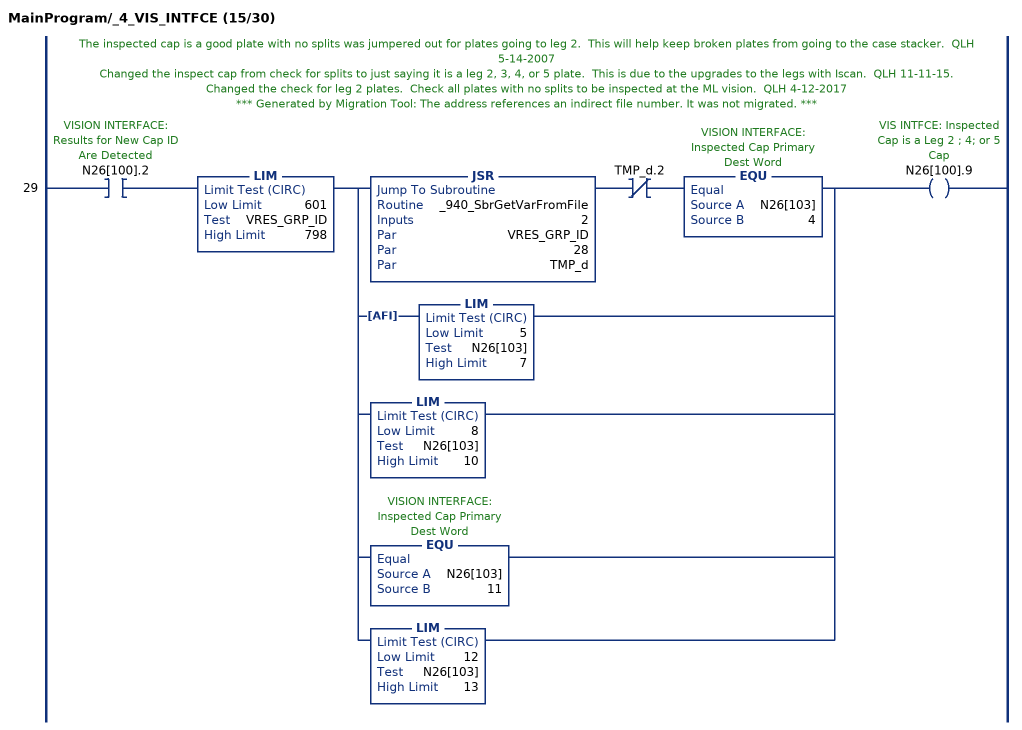
   // The inspected cap is a good plate with no splits was jumpered out for plates going to leg 2.  This will help keep broken plates from going to the case stacker.  QLH 5-14-2007
   // Changed the inspect cap from check for splits to just saying it is a leg 2, 3, 4, or 5 plate.  This is due to the upgrades to the legs with Iscan.  QLH 11-11-15.  Changed the check for leg 2 plates.  Check all plates with no splits to be inspected at the ML vision.  QLH 4-12-2017
   // *** Generated by Migration Tool: The address references an indirect file number. It was not migrated. ***
   29: XIC(N26[100].2)LIM(601,VRES_GRP_ID,798)[JSR(_940_SbrGetVarFromFile,2,VRES_GRP_ID,28,TMP_d) XIO(TMP_d.2) EQU(N26[103],4) ,AFI() LIM(5,N26[103],7) ,LIM(8,N26[103],10) ,EQU(N26[103],11) ,LIM(12,N26[103],13) ]OTE(N26[100].9);
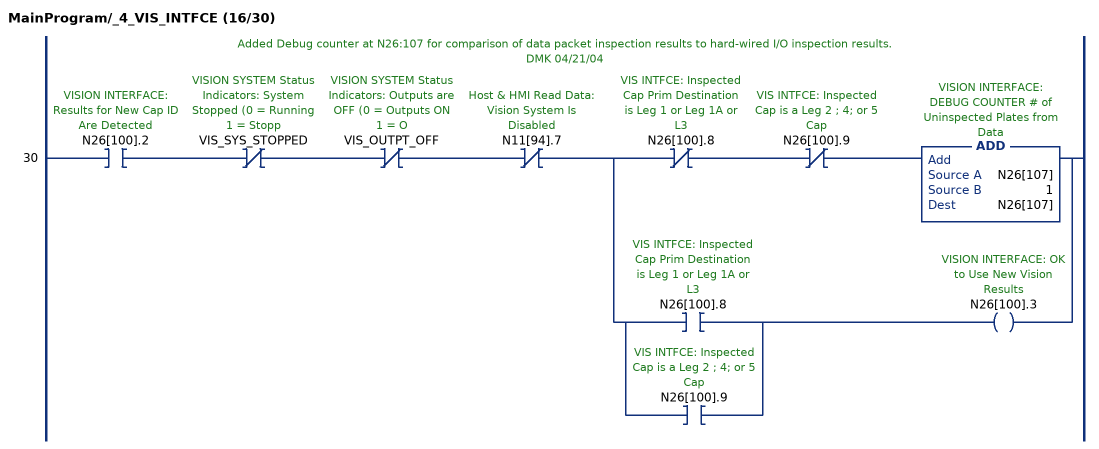
   // Added Debug counter at N26:107 for comparison of data packet inspection results to hard-wired I/O inspection results.
   // DMK 04/21/04
   30: XIC(N26[100].2)XIO(VIS_SYS_STOPPED)XIO(VIS_OUTPT_OFF)XIO(N11[94].7)[XIO(N26[100].8) XIO(N26[100].9) ADD(N26[107],1,N26[107]) ,[XIC(N26[100].8) ,XIC(N26[100].9) ] OTE(N26[100].3) ];
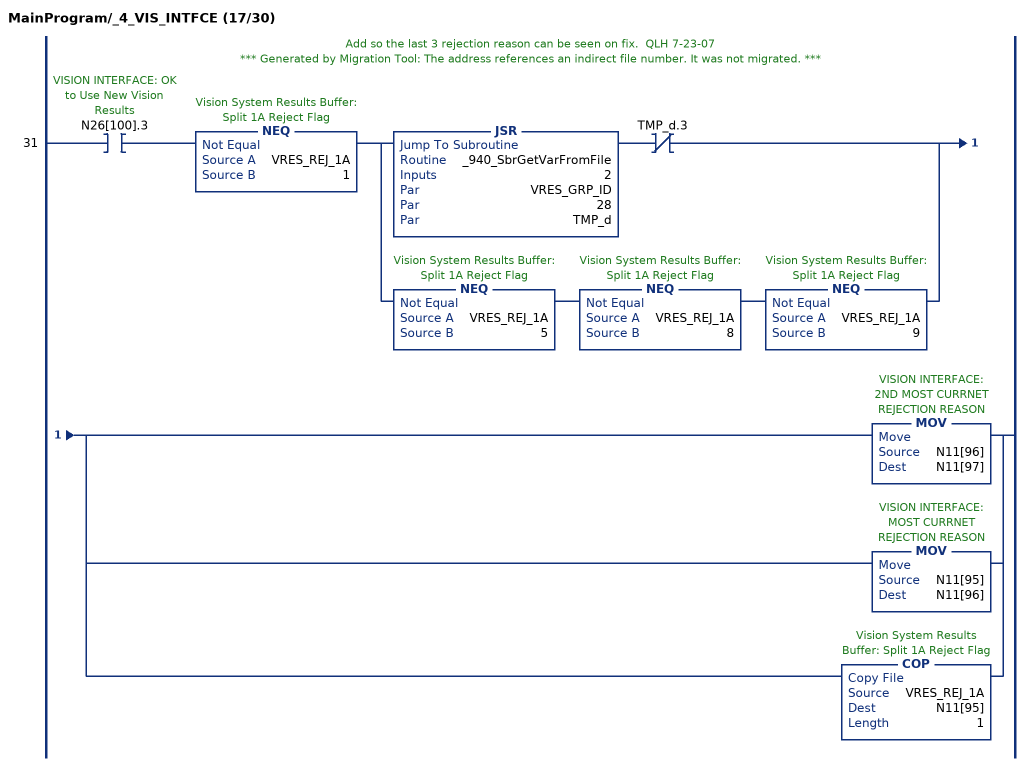
   // Add so the last 3 rejection reason can be seen on fix.  QLH 7-23-07
   // *** Generated by Migration Tool: The address references an indirect file number. It was not migrated. ***
   31: XIC(N26[100].3)NEQ(VRES_REJ_1A,1)[JSR(_940_SbrGetVarFromFile,2,VRES_GRP_ID,28,TMP_d) XIO(TMP_d.3) ,NEQ(VRES_REJ_1A,5) NEQ(VRES_REJ_1A,8) NEQ(VRES_REJ_1A,9) ][MOV(N11[96],N11[97]) ,MOV(N11[95],N11[96]) ,COP(VRES_REJ_1A,N11[95],1) ];
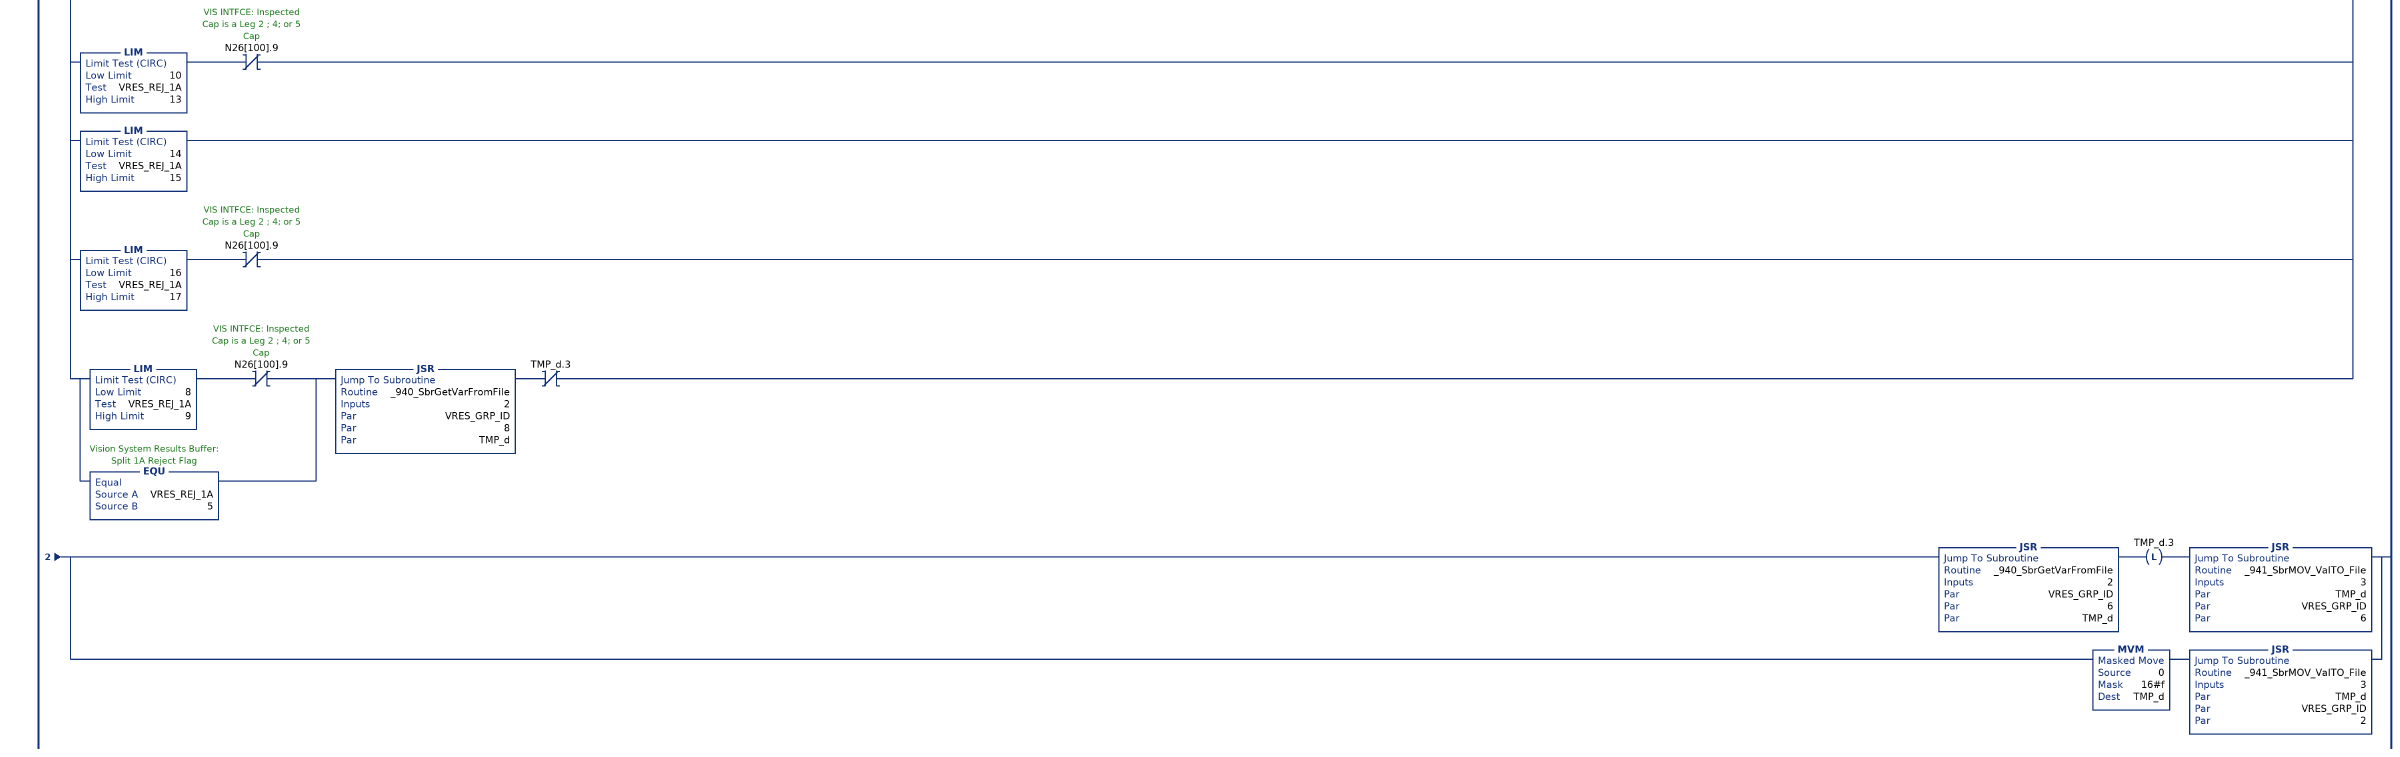
   // Will not look at width errors on 1/2 inch 2 plate splits for Leg 2.  They are keeping trim on the plate to help with a size they are cutting.  Will take out once run is complete.  QLH 5/12/10 Same change 7-2-10 QLH same 3/10/11 QLH
   // *** Generated by Migration Tool: The address references an indirect file number. It was not migrated. ***
   // *** Generated by Migration Tool: The address references an indirect file number. It was not migrated. ***
   // *** Generated by Migration Tool: The address references an indirect file number. It was not migrated. ***
   // *** Generated by Migration Tool: The address references an indirect file number. It was not migrated. ***
   // *** Generated by Migration Tool: The address references an indirect file number. It was not migrated. ***
   // *** Generated by Migration Tool: The address references an indirect file number. It was not migrated. ***
   // *** Generated by Migration Tool: The address references an indirect file number. It was not migrated. ***
   // *** Generated by Migration Tool: The address references an indirect file number. It was not migrated. ***
   // *** Generated by Migration Tool: The address references an indirect file number. It was not migrated. ***
   // *** Generated by Migration Tool: The address references an indirect file number. It was not migrated. ***
   32: XIC(N26[100].3)[[LIM(2,VRES_REJ_1A,3) XIO(N26[100].9) ,EQU(VRES_REJ_1A,4) ,LIM(6,VRES_REJ_1A,7) XIO(N26[100].9) [LIM(601,VRES_GRP_ID,798) JSR(_940_SbrGetVarFromFile,2,VRES_GRP_ID,28,TMP_d) XIC(TMP_d.2) ,NEQ(N26[99],4) ,LIM(601,VRES_GRP_ID,798) JSR(_940_SbrGetVarFromFile,2,VRES_GRP_ID,8,TMP_d) NEQ(TMP_d,6912) JSR(_940_SbrGetVarFromFile,2,VRES_GRP_ID,10,TMP_d) NEQ(TMP_d,6912) JSR(_940_SbrGetVarFromFile,2,VRES_GRP_ID,8,TMP_d) NEQ(TMP_d,6528) JSR(_940_SbrGetVarFromFile,2,VRES_GRP_ID,10,TMP_d) NEQ(TMP_d,6528) JSR(_940_SbrGetVarFromFile,2,VRES_GRP_ID,8,TMP_d) NEQ(TMP_d,6400) JSR(_940_SbrGetVarFromFile,2,VRES_GRP_ID,10,TMP_d) NEQ(TMP_d,6400) ,XIO(xAlwaysOFF) ] ,LIM(10,VRES_REJ_1A,13) XIO(N26[100].9) ,LIM(14,VRES_REJ_1A,15) ,LIM(16,VRES_REJ_1A,17) XIO(N26[100].9) ] ,[LIM(8,VRES_REJ_1A,9) XIO(N26[100].9) ,EQU(VRES_REJ_1A,5) ] JSR(_940_SbrGetVarFromFile,2,VRES_GRP_ID,8,TMP_d) XIO(TMP_d.3) ][JSR(_940_SbrGetVarFromFile,2,VRES_GRP_ID,6,TMP_d) OTL(TMP_d.3) JSR(_941_SbrMOV_ValTO_File,3,TMP_d,VRES_GRP_ID,6) ,MVM(0,16#f,TMP_d) JSR(_941_SbrMOV_ValTO_File,3,TMP_d,VRES_GRP_ID,2) ];
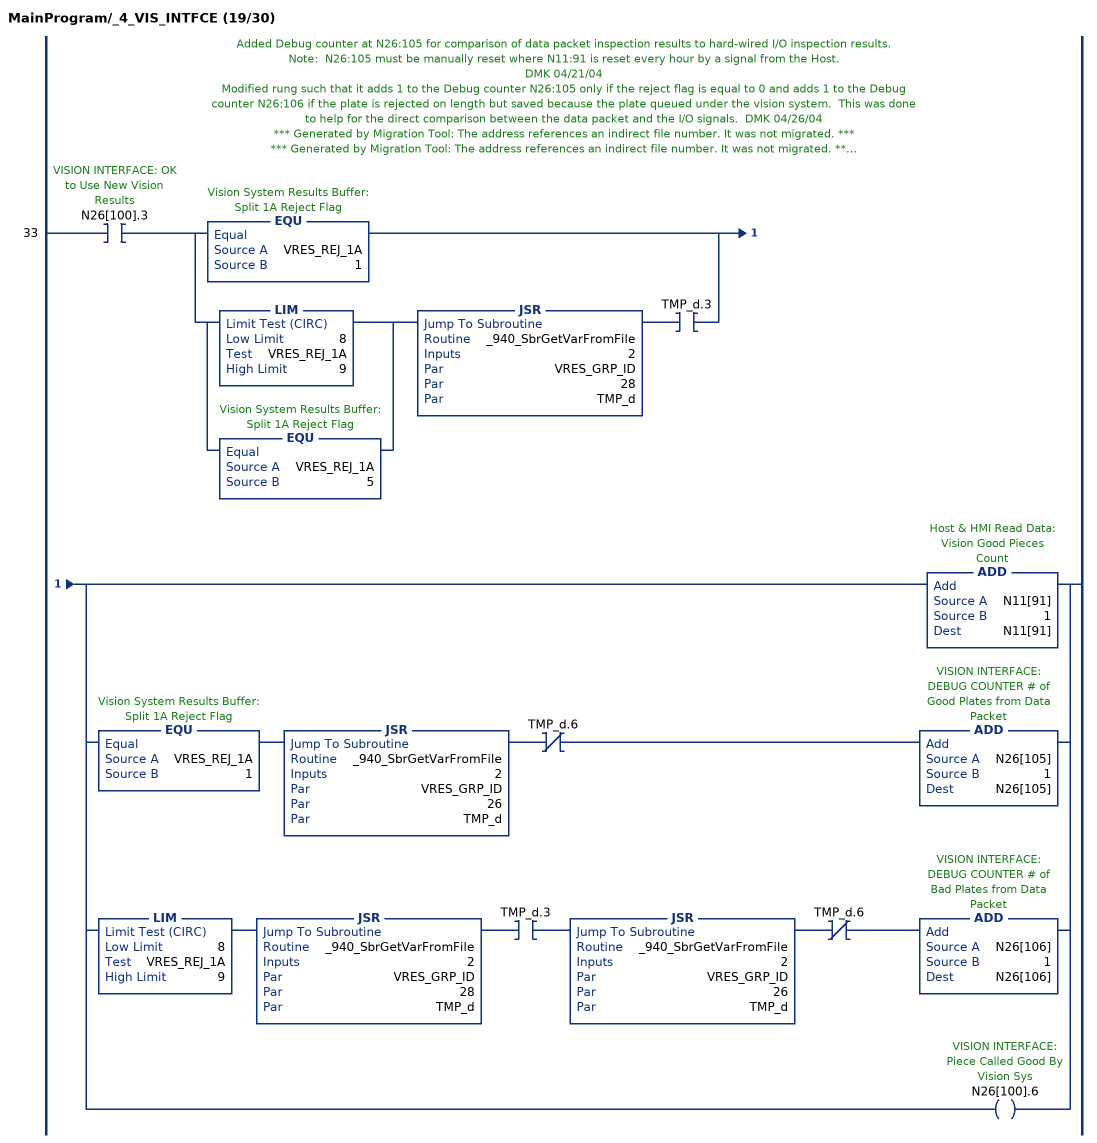
   // Added Debug counter at N26:105 for comparison of data packet inspection results to hard-wired I/O inspection results.
   // Note:  N26:105 must be manually reset where N11:91 is reset every hour by a signal from the Host.
   // DMK 04/21/04
   // Modified rung such that it adds 1 to the Debug counter N26:105 only if the reject flag is equal to 0 and adds 1 to the Debug
   // counter N26:106 if the plate is rejected on length but saved because the plate queued under the vision system.  This was done
   // to help for the direct comparison between the data packet and the I/O signals.  DMK 04/26/04
   // *** Generated by Migration Tool: The address references an indirect file number. It was not migrated. ***
   // *** Generated by Migration Tool: The address references an indirect file number. It was not migrated. ***
   // *** Generated by Migration Tool: The address references an indirect file number. It was not migrated. ***
   // *** Generated by Migration Tool: The address references an indirect file number. It was not migrated. ***
   33: XIC(N26[100].3)[EQU(VRES_REJ_1A,1) ,[LIM(8,VRES_REJ_1A,9) ,EQU(VRES_REJ_1A,5) ] JSR(_940_SbrGetVarFromFile,2,VRES_GRP_ID,28,TMP_d) XIC(TMP_d.3) ][ADD(N11[91],1,N11[91]) ,EQU(VRES_REJ_1A,1) JSR(_940_SbrGetVarFromFile,2,VRES_GRP_ID,26,TMP_d) XIO(TMP_d.6) ADD(N26[105],1,N26[105]) ,LIM(8,VRES_REJ_1A,9) JSR(_940_SbrGetVarFromFile,2,VRES_GRP_ID,28,TMP_d) XIC(TMP_d.3) JSR(_940_SbrGetVarFromFile,2,VRES_GRP_ID,26,TMP_d) XIO(TMP_d.6) ADD(N26[106],1,N26[106]) ,OTE(N26[100].6) ];
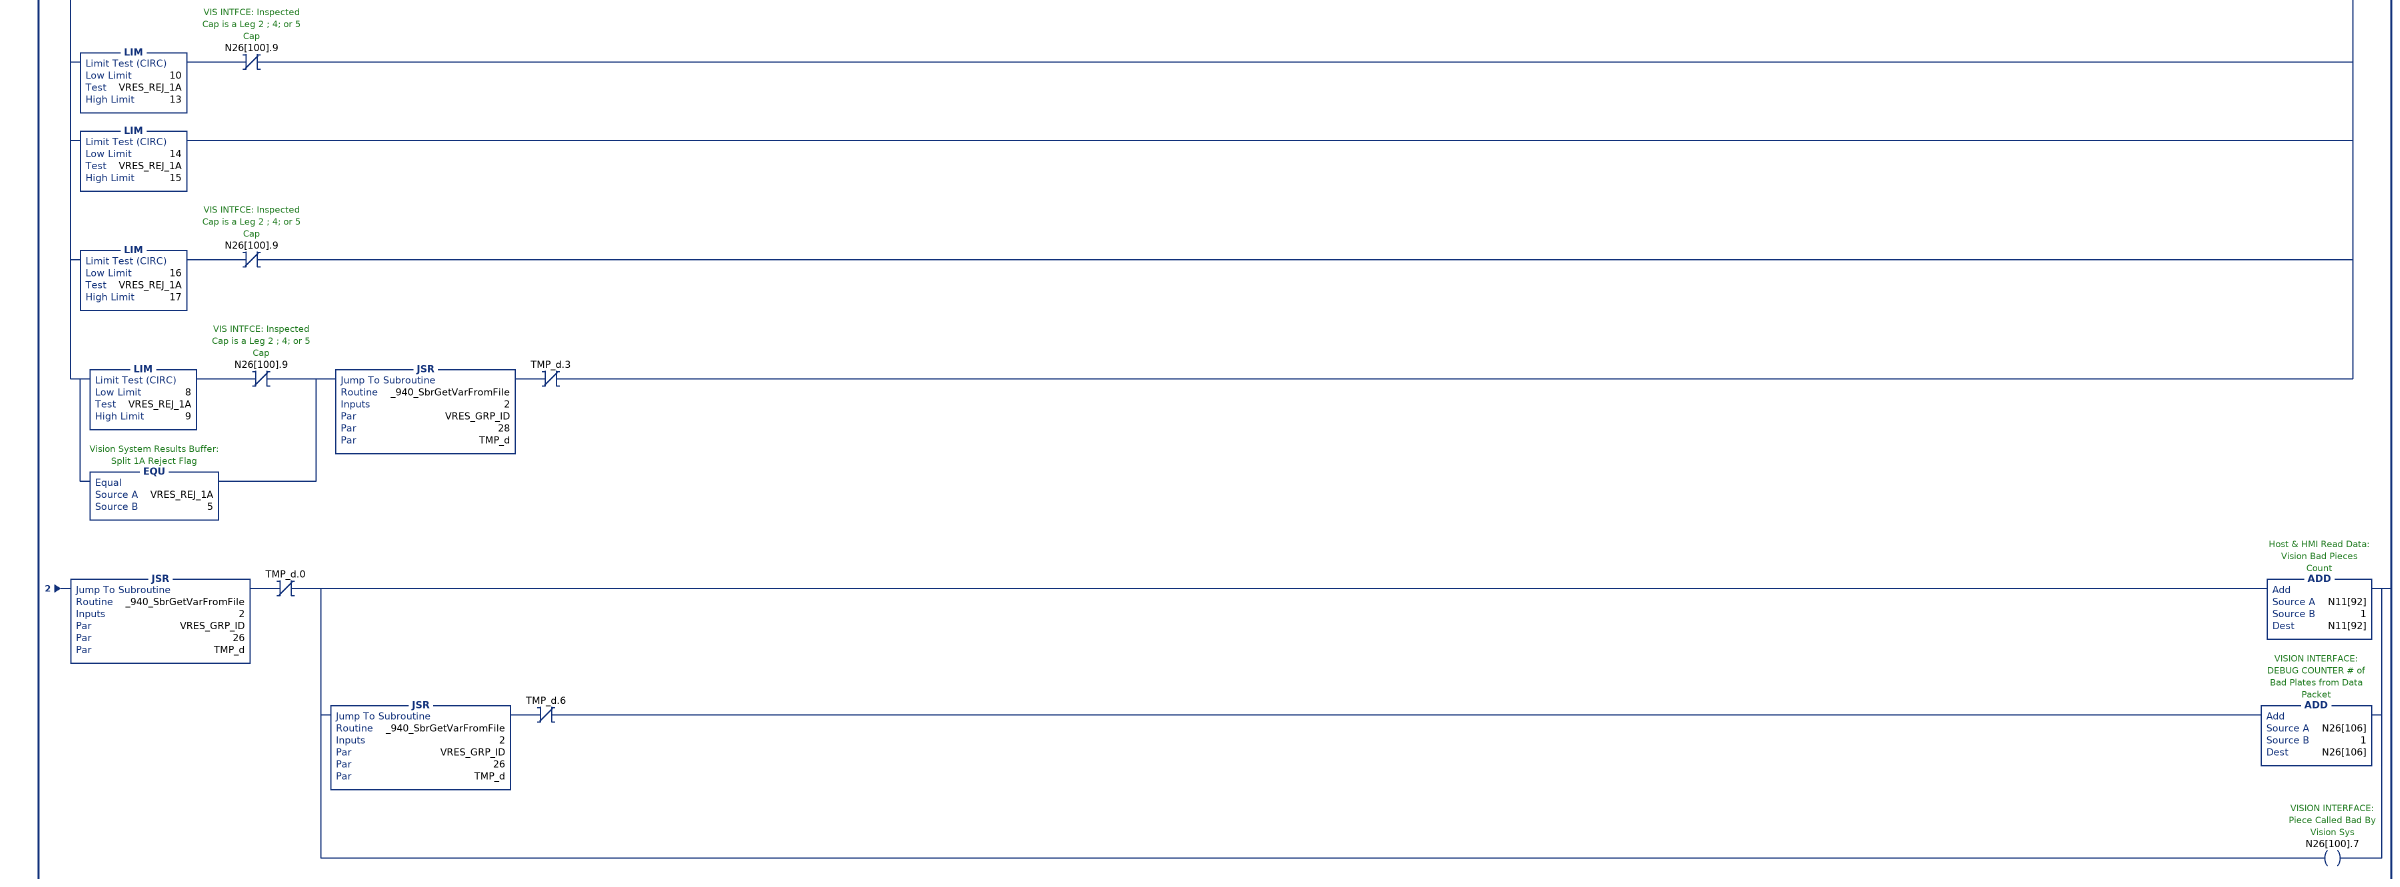
   // Added Debug counter at N26:106 for comparison of data packet inspection results to hard-wired I/O inspection results.
   // Note:  N26:106 must be manually reset where N11:92 is reset every hour by a signal from the Host.
   // DMK 04/21/04
   // Will not look at width errors on 1/2 inch 2 plate splits for Leg 2.  They are keeping trim on the plate to help with a size they are cutting.  Will take out once run is complete.  QLH 5/12/10
   // *** Generated by Migration Tool: The address references an indirect file number. It was not migrated. ***
   // *** Generated by Migration Tool: The address references an indirect file number. It was not migrated. ***
   // *** Generated by Migration Tool: The address references an indirect file number. It was not migrated. ***
   // *** Generated by Migration Tool: The address references an indirect file number. It was not migrated. ***
   // *** Generated by Migration Tool: The address references an indirect file number. It was not migrated. ***
   // *** Generated by Migration Tool: The address references an indirect file number. It was not migrated. ***
   // *** Generated by Migration Tool: The address references an indirect file number. It was not migrated. ***
   // *** Generated by Migration Tool: The address references an indirect file number. It was not migrated. ***
   // *** Generated by Migration Tool: The address references an indirect file number. It was not migrated. ***
   // *** Generated by Migration Tool: The address references an indirect file number. It was not migrated. ***
   34: XIC(N26[100].3)[[LIM(2,VRES_REJ_1A,3) XIO(N26[100].9) ,EQU(VRES_REJ_1A,4) ,LIM(6,VRES_REJ_1A,7) XIO(N26[100].9) [LIM(601,VRES_GRP_ID,798) JSR(_940_SbrGetVarFromFile,2,VRES_GRP_ID,28,TMP_d) XIC(TMP_d.2) ,NEQ(N26[99],4) ,LIM(601,VRES_GRP_ID,798) JSR(_940_SbrGetVarFromFile,2,VRES_GRP_ID,8,TMP_d) NEQ(TMP_d,6912) JSR(_940_SbrGetVarFromFile,2,VRES_GRP_ID,10,TMP_d) NEQ(TMP_d,6912) JSR(_940_SbrGetVarFromFile,2,VRES_GRP_ID,8,TMP_d) NEQ(TMP_d,6528) JSR(_940_SbrGetVarFromFile,2,VRES_GRP_ID,10,TMP_d) NEQ(TMP_d,6528) JSR(_940_SbrGetVarFromFile,2,VRES_GRP_ID,8,TMP_d) NEQ(TMP_d,6400) JSR(_940_SbrGetVarFromFile,2,VRES_GRP_ID,10,TMP_d) NEQ(TMP_d,6400) ,XIO(xAlwaysOFF) ] ,LIM(10,VRES_REJ_1A,13) XIO(N26[100].9) ,LIM(14,VRES_REJ_1A,15) ,LIM(16,VRES_REJ_1A,17) XIO(N26[100].9) ] ,[LIM(8,VRES_REJ_1A,9) XIO(N26[100].9) ,EQU(VRES_REJ_1A,5) ] JSR(_940_SbrGetVarFromFile,2,VRES_GRP_ID,28,TMP_d) XIO(TMP_d.3) ]JSR(_940_SbrGetVarFromFile,2,VRES_GRP_ID,26,TMP_d)XIO(TMP_d.0)[ADD(N11[92],1,N11[92]) ,JSR(_940_SbrGetVarFromFile,2,VRES_GRP_ID,26,TMP_d) XIO(TMP_d.6) ADD(N26[106],1,N26[106]) ,OTE(N26[100].7) ];
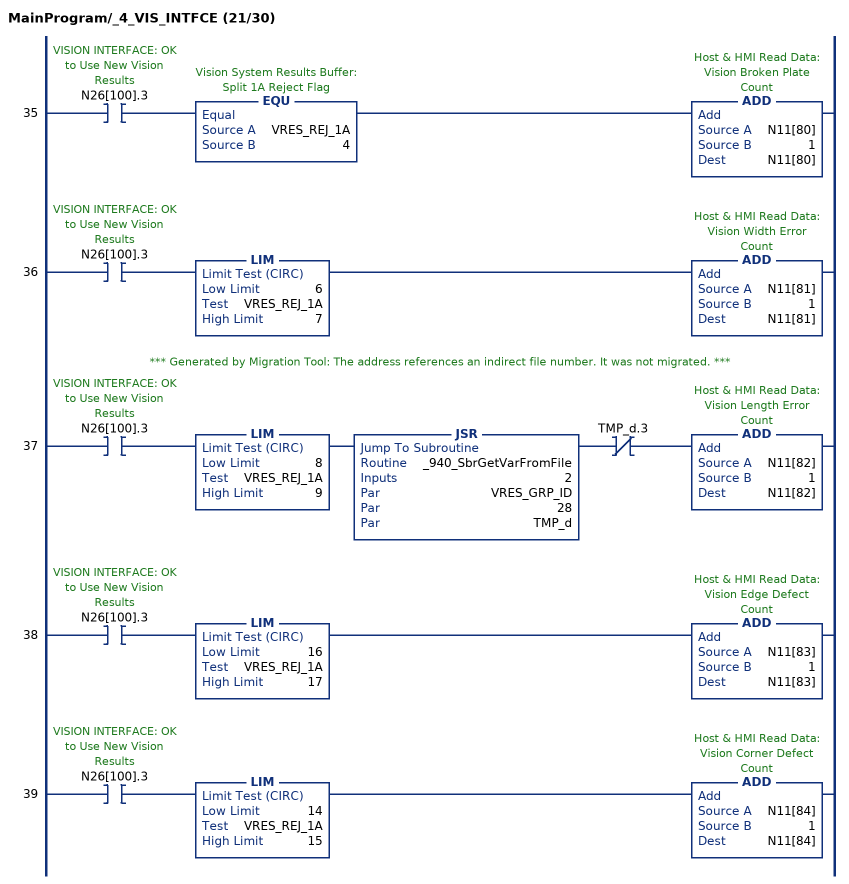
   35: XIC(N26[100].3)EQU(VRES_REJ_1A,4)ADD(N11[80],1,N11[80]);
   36: XIC(N26[100].3)LIM(6,VRES_REJ_1A,7)ADD(N11[81],1,N11[81]);
   // *** Generated by Migration Tool: The address references an indirect file number. It was not migrated. ***
   37: XIC(N26[100].3)LIM(8,VRES_REJ_1A,9)JSR(_940_SbrGetVarFromFile,2,VRES_GRP_ID,28,TMP_d)XIO(TMP_d.3)ADD(N11[82],1,N11[82]);
   38: XIC(N26[100].3)LIM(16,VRES_REJ_1A,17)ADD(N11[83],1,N11[83]);
   39: XIC(N26[100].3)LIM(14,VRES_REJ_1A,15)ADD(N11[84],1,N11[84]);
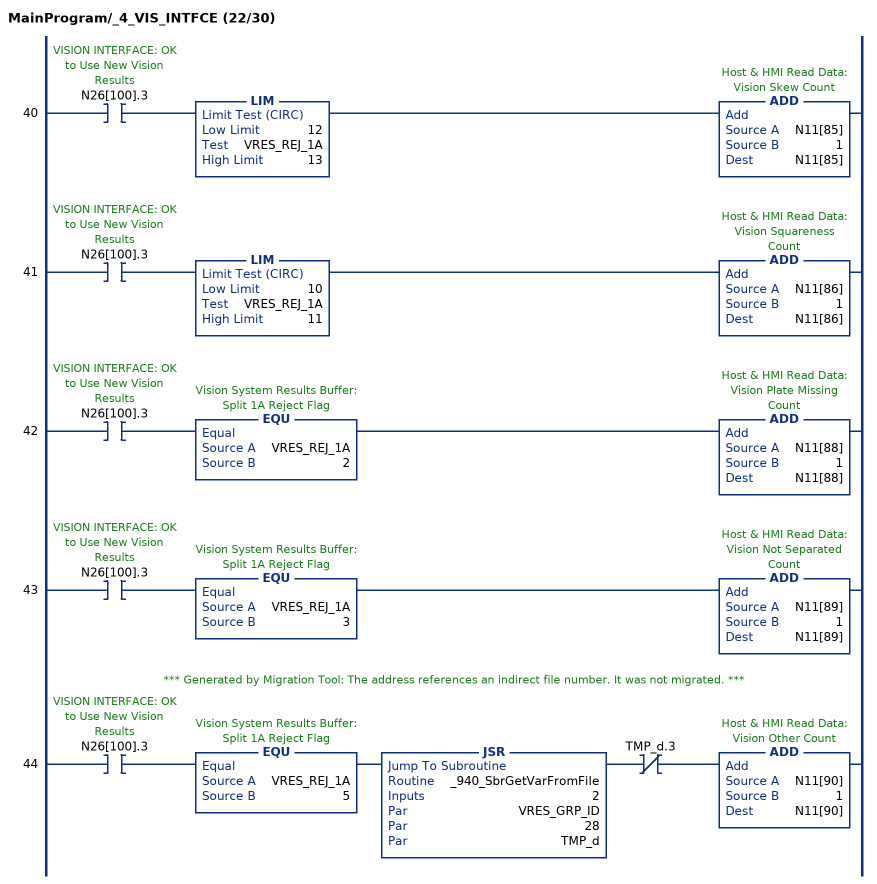
   40: XIC(N26[100].3)LIM(12,VRES_REJ_1A,13)ADD(N11[85],1,N11[85]);
   41: XIC(N26[100].3)LIM(10,VRES_REJ_1A,11)ADD(N11[86],1,N11[86]);
   42: XIC(N26[100].3)EQU(VRES_REJ_1A,2)ADD(N11[88],1,N11[88]);
   43: XIC(N26[100].3)EQU(VRES_REJ_1A,3)ADD(N11[89],1,N11[89]);
   // *** Generated by Migration Tool: The address references an indirect file number. It was not migrated. ***
   44: XIC(N26[100].3)EQU(VRES_REJ_1A,5)JSR(_940_SbrGetVarFromFile,2,VRES_GRP_ID,28,TMP_d)XIO(TMP_d.3)ADD(N11[90],1,N11[90]);
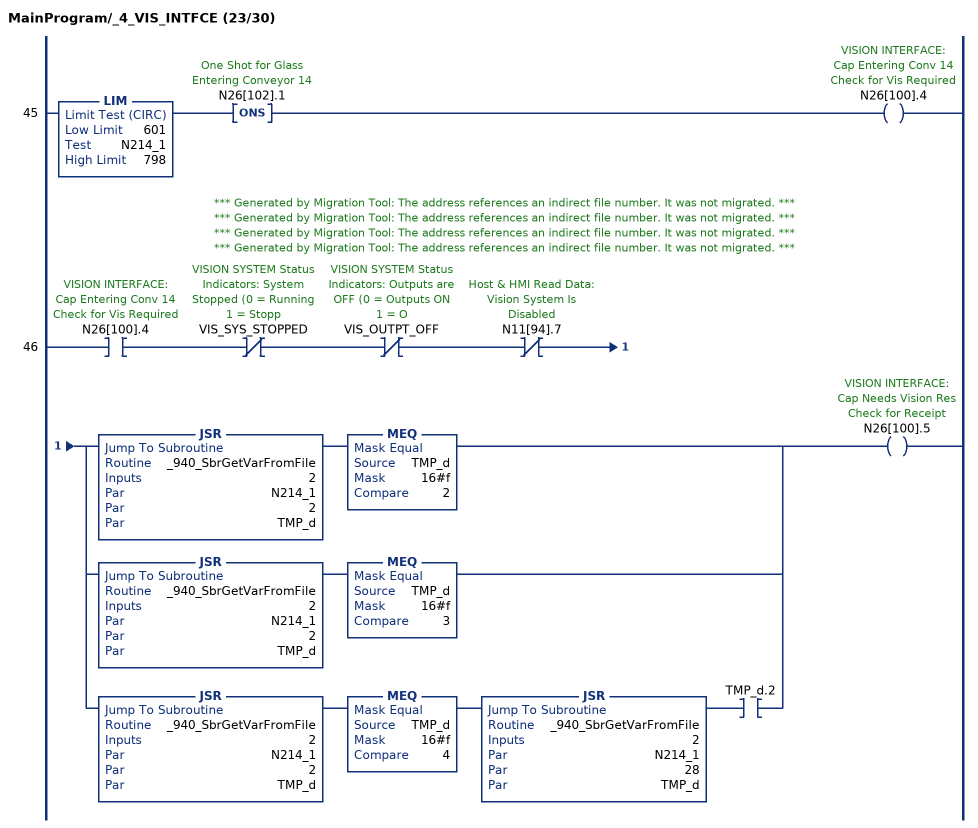
   45: LIM(601,N214_1,798)ONS(N26[102].1)OTE(N26[100].4);
   // *** Generated by Migration Tool: The address references an indirect file number. It was not migrated. ***
   // *** Generated by Migration Tool: The address references an indirect file number. It was not migrated. ***
   // *** Generated by Migration Tool: The address references an indirect file number. It was not migrated. ***
   // *** Generated by Migration Tool: The address references an indirect file number. It was not migrated. ***
   46: XIC(N26[100].4)XIO(VIS_SYS_STOPPED)XIO(VIS_OUTPT_OFF)XIO(N11[94].7)[JSR(_940_SbrGetVarFromFile,2,N214_1,2,TMP_d) MEQ(TMP_d,16#f,2) ,JSR(_940_SbrGetVarFromFile,2,N214_1,2,TMP_d) MEQ(TMP_d,16#f,3) ,JSR(_940_SbrGetVarFromFile,2,N214_1,2,TMP_d) MEQ(TMP_d,16#f,4) JSR(_940_SbrGetVarFromFile,2,N214_1,28,TMP_d) XIC(TMP_d.2) ]OTE(N26[100].5);
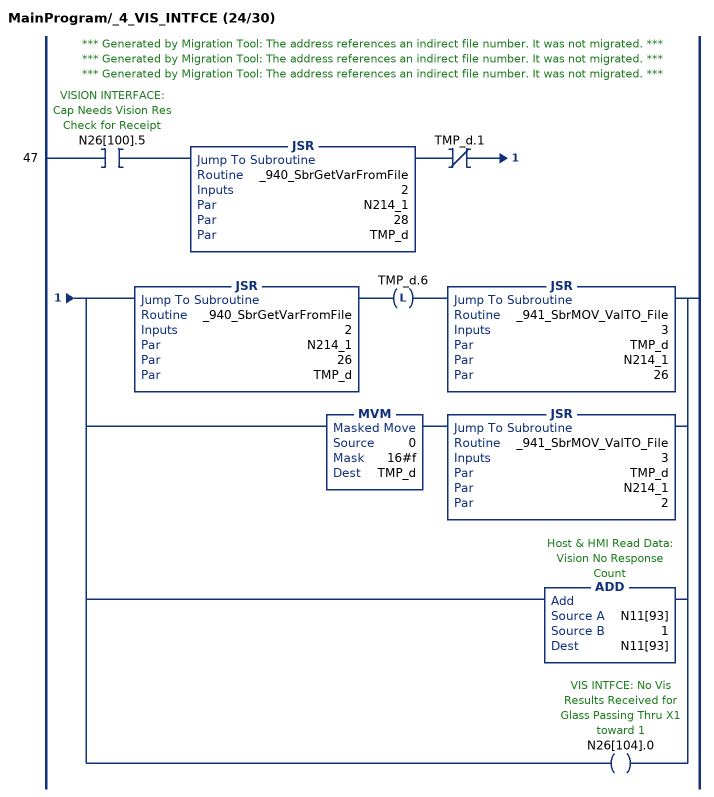
   // *** Generated by Migration Tool: The address references an indirect file number. It was not migrated. ***
   // *** Generated by Migration Tool: The address references an indirect file number. It was not migrated. ***
   // *** Generated by Migration Tool: The address references an indirect file number. It was not migrated. ***
   47: XIC(N26[100].5)JSR(_940_SbrGetVarFromFile,2,N214_1,28,TMP_d)XIO(TMP_d.1)[JSR(_940_SbrGetVarFromFile,2,N214_1,26,TMP_d) OTL(TMP_d.6) JSR(_941_SbrMOV_ValTO_File,3,TMP_d,N214_1,26) ,MVM(0,16#f,TMP_d) JSR(_941_SbrMOV_ValTO_File,3,TMP_d,N214_1,2) ,ADD(N11[93],1,N11[93]) ,OTE(N26[104].0) ];
